HMI tags "Sim Stations"
   "HMI Data: Warehouse HMI_simStations_down" : Push Button Data = PLC "HMI Data: Warehouse HMI".simStations.down, 100 ms
   "HMI Data: Warehouse HMI_simStations_me{0}" : Station: Sim Data = PLC "HMI Data: Warehouse HMI".simStations.me[0] AT %DB1.DBX0.0, 100 ms
   "HMI Data: Warehouse HMI_simStations_me{1}" : Station: Sim Data = PLC "HMI Data: Warehouse HMI".simStations.me[1], 100 ms
   "HMI Data: Warehouse HMI_simStations_me{10}" : Station: Sim Data = PLC "HMI Data: Warehouse HMI".simStations.me[10], 100 ms
   "HMI Data: Warehouse HMI_simStations_me{11}" : Station: Sim Data = PLC "HMI Data: Warehouse HMI".simStations.me[11], 100 ms
   "HMI Data: Warehouse HMI_simStations_me{2}" : Station: Sim Data = PLC "HMI Data: Warehouse HMI".simStations.me[2], 100 ms
   "HMI Data: Warehouse HMI_simStations_me{3}" : Station: Sim Data = PLC "HMI Data: Warehouse HMI".simStations.me[3], 100 ms
   "HMI Data: Warehouse HMI_simStations_me{4}" : Station: Sim Data = PLC "HMI Data: Warehouse HMI".simStations.me[4], 100 ms
   "HMI Data: Warehouse HMI_simStations_me{5}" : Station: Sim Data = PLC "HMI Data: Warehouse HMI".simStations.me[5], 100 ms
   "HMI Data: Warehouse HMI_simStations_me{6}" : Station: Sim Data = PLC "HMI Data: Warehouse HMI".simStations.me[6], 100 ms
   "HMI Data: Warehouse HMI_simStations_me{7}" : Station: Sim Data = PLC "HMI Data: Warehouse HMI".simStations.me[7], 100 ms
   "HMI Data: Warehouse HMI_simStations_me{8}" : Station: Sim Data = PLC "HMI Data: Warehouse HMI".simStations.me[8], 100 ms
   "HMI Data: Warehouse HMI_simStations_me{9}" : Station: Sim Data = PLC "HMI Data: Warehouse HMI".simStations.me[9], 100 ms
   "HMI Data: Warehouse HMI_simStations_up" : Push Button Data = PLC "HMI Data: Warehouse HMI".simStations.up, 100 ms

HMI tags "Settings: Interface"
   "HMI Data: Warehouse HMI_settings_assign" : Push Button Data = PLC "HMI Data: Warehouse HMI".settings.assign, 100 ms
   "HMI Data: Warehouse HMI_settings_partNumber" : Part_Number_Double.UDT = PLC "HMI Data: Warehouse HMI".settings.partNumber, 100 ms
   "HMI Data: Warehouse HMI_settings_critical" : IO Field Data: Label with Data = PLC "HMI Data: Warehouse HMI".settings.critical, 100 ms
   "HMI Data: Warehouse HMI_settings_total" : IO Field Data: Label with Data = PLC "HMI Data: Warehouse HMI".settings.total, 100 ms
   "HMI Data: Warehouse HMI_settings_dropzone" : IO Field Data: Label with Data = PLC "HMI Data: Warehouse HMI".settings.dropzone, 100 ms
   "HMI Data: Warehouse HMI_settings_line" : IO Field Data: Label with Data = PLC "HMI Data: Warehouse HMI".settings.line, 100 ms
   "HMI Data: Warehouse HMI_settings_selectButton" : Push Button Data = PLC "HMI Data: Warehouse HMI".settings.selectButton, 100 ms
   "HMI Data: Warehouse HMI_settings_selectWip" : Push Button Data = PLC "HMI Data: Warehouse HMI".settings.selectWip, 100 ms
   "HMI Data: Warehouse HMI_settings_selectStation" : Push Button Data = PLC "HMI Data: Warehouse HMI".settings.selectStation, 100 ms
   "HMI Data: Warehouse HMI_settings_stnTableNavBar_hmi" : Nav Bar Data: HMI = PLC "HMI Data: Warehouse HMI".settings.stnTableNavBar.hmi AT %DB1.DBW0, 100 ms

HMI tags "Settings: Feedback"
   "HMI Data: Warehouse HMI_settings_stationRows{0}" : Settings Station Row Data = PLC "HMI Data: Warehouse HMI".settings.stationRows[0], 100 ms
   "HMI Data: Warehouse HMI_settings_stationRows{1}" : Settings Station Row Data = PLC "HMI Data: Warehouse HMI".settings.stationRows[1], 100 ms
   "HMI Data: Warehouse HMI_settings_stationRows{2}" : Settings Station Row Data = PLC "HMI Data: Warehouse HMI".settings.stationRows[2], 100 ms

graphic list "Vertical Table Nav Bar": 0 '100 x 100 Top'; 1 '100 x 100 Actuated Top'; 2 '100 x 100 Page Up'; 3 '100 x 100 Actuated Page Up'; 4 '100 x 100 Line Up'; 5 '100 x 100 Actuated Line Up'; 6 '100 x 100 Line Down'; 7 '100 x 100 Actuated Line Down'; 8 '100 x 100 Page Down'; 9 '100 x 100 Actuated Page Down'; 10 '100 x 100 Bottom'; 11 '100 x 100 Actuated Bottom'

screen "1 PART CALL" 1366x768
   on GenerateScreen: SetTag("HMI Data: Warehouse HMI_screenNumber", 1)
   Rectangle "Settings Tab Background" at 682,0 size 684x68
      Appearance <- "HMI Data: Warehouse HMI_screenNumber"
   Rectangle "Part Call Tab Background" at 0,0 size 685x68
      Appearance <- "HMI Data: Warehouse HMI_screenNumber"
   Rectangle "Settings Tab Border Hide" at 685,61 size 678x20
      Visibility <- "HMI Data: Warehouse HMI_screenNumber"
   Rectangle "Part Call Tab Border Hide" at 3,61 size 679x20
      Visibility <- "HMI Data: Warehouse HMI_screenNumber"
   Button "Settings Screen" at 683,0 size 683x68; TextOff 'SETTINGS'; Authorization "User administration"
      on Release: ActivateScreen("2 SETTINGS", 0)
   Button "Part Call Screen" at 0,0 size 683x68; TextOff 'PART CALL'
      on Release: ActivateScreen("1 PART CALL", 0)
   TextField "Header Line" at 32,112 size 216x53; Text 'LINE'
   TextField "Header Drop Zone" at 238,112 size 236x53; Text 'DROP ZONE'
   TextField "Header Part Number" at 474,112 size 648x53; Text 'PART NUMBER'
   TextField "Header Time" at 1112,112 size 222x53; Text 'TIME'
   ScreenModuleView "TableRow00" at 27,170 size 1312x52; ScreenModuleType ""
      Guid_{11997190-27688} <- "HMI Data: Warehouse HMI_partCall_row{0}"
      on Guid_{11997190-83214}: ActivateScreen("3 BARCODE", 0)
   ScreenModuleView "TableRow01" at 27,222 size 1312x52; ScreenModuleType ""
      Guid_{11997190-27688} <- "HMI Data: Warehouse HMI_partCall_row{1}"
      on Guid_{11997190-83214}: ActivateScreen("3 BARCODE", 0)
   ScreenModuleView "TableRow02" at 27,274 size 1312x52; ScreenModuleType ""
      Guid_{11997190-27688} <- "HMI Data: Warehouse HMI_partCall_row{2}"
      on Guid_{11997190-83214}: ActivateScreen("3 BARCODE", 0)
   ScreenModuleView "TableRow03" at 27,326 size 1312x52; ScreenModuleType ""
      Guid_{11997190-27688} <- "HMI Data: Warehouse HMI_partCall_row{3}"
      on Guid_{11997190-83214}: ActivateScreen("3 BARCODE", 0)
   ScreenModuleView "TableRow04" at 27,378 size 1312x52; ScreenModuleType ""
      Guid_{11997190-27688} <- "HMI Data: Warehouse HMI_partCall_row{4}"
      on Guid_{11997190-83214}: ActivateScreen("3 BARCODE", 0)
   ScreenModuleView "TableRow05" at 27,430 size 1312x52; ScreenModuleType ""
      Guid_{11997190-27688} <- "HMI Data: Warehouse HMI_partCall_row{5}"
      on Guid_{11997190-83214}: ActivateScreen("3 BARCODE", 0)
   ScreenModuleView "TableRow06" at 27,482 size 1312x52; ScreenModuleType ""
      Guid_{11997190-27688} <- "HMI Data: Warehouse HMI_partCall_row{6}"
      on Guid_{11997190-83214}: ActivateScreen("3 BARCODE", 0)
   ScreenModuleView "TableRow07" at 27,534 size 1312x52; ScreenModuleType ""
      Guid_{11997190-27688} <- "HMI Data: Warehouse HMI_partCall_row{7}"
      on Guid_{11997190-83214}: ActivateScreen("3 BARCODE", 0)
   ScreenModuleView "TableRow08" at 27,586 size 1312x52; ScreenModuleType ""
      Guid_{11997190-27688} <- "HMI Data: Warehouse HMI_partCall_row{8}"
      on Guid_{11997190-83214}: ActivateScreen("3 BARCODE", 0)
   ScreenModuleView "TableRow09" at 27,638 size 1312x52; ScreenModuleType ""
      Guid_{11997190-27688} <- "HMI Data: Warehouse HMI_partCall_row{9}"
      on Guid_{11997190-83214}: ActivateScreen("3 BARCODE", 0)
   ScreenModuleView "TableRow10" at 27,690 size 1312x52; ScreenModuleType ""
      Guid_{11997190-27688} <- "HMI Data: Warehouse HMI_partCall_row{10}"
      on Guid_{11997190-83214}: ActivateScreen("3 BARCODE", 0)

SlideinScreen "GraphX_Slidein_Bottom" 1366x80
   ScreenModuleView "Top" at 0,0 size 227x80; Guid_{11997190-63799} "Top"; ScreenModuleType ""
      Guid_{11997190-63779} <- "HMI Data: Warehouse HMI_tableNav_top"
   ScreenModuleView "Page Up" at 227,0 size 228x80; Guid_{11997190-63799} "pageUp"; ScreenModuleType ""
      Guid_{11997190-63779} <- "HMI Data: Warehouse HMI_tableNav_pageUp"
   ScreenModuleView "Line Up" at 455,0 size 228x80; Guid_{11997190-63799} "Up"; ScreenModuleType ""
      Guid_{11997190-63779} <- "HMI Data: Warehouse HMI_tableNav_lineUp"
   ScreenModuleView "Line Down" at 683,0 size 228x80; Guid_{11997190-63799} "Down"; ScreenModuleType ""
      Guid_{11997190-63779} <- "HMI Data: Warehouse HMI_tableNav_lineDown"
   ScreenModuleView "Page Down" at 911,0 size 228x80; Guid_{11997190-63799} "PageDown"; ScreenModuleType ""
      Guid_{11997190-63779} <- "HMI Data: Warehouse HMI_tableNav_pageDown"
   ScreenModuleView "Bottom" at 1138,0 size 228x80; Guid_{11997190-63799} "Bottom"; ScreenModuleType ""
      Guid_{11997190-63779} <- "HMI Data: Warehouse HMI_tableNav_bottom"
   TextField "Text field_1" at 0,0 size 1366x80; Text 'NOT USED'
      Visibility <- "HMI Data: Warehouse HMI_screenNumber"

SlideinScreen "GraphX_Slidein_Right" 449x768
   ScreenModuleView "Station Sim_1" at 5,5 size 106x232; ScreenModuleType ""
      Guid_{11997190-89108} <- "HMI Data: Warehouse HMI_simStations_me{0}"
   ScreenModuleView "Station Sim_2" at 116,5 size 106x232; ScreenModuleType ""
      Guid_{11997190-89108} <- "HMI Data: Warehouse HMI_simStations_me{1}"
   ScreenModuleView "Station Sim_3" at 227,5 size 106x232; ScreenModuleType ""
      Guid_{11997190-89108} <- "HMI Data: Warehouse HMI_simStations_me{2}"
   ScreenModuleView "Station Sim_4" at 338,5 size 106x232; ScreenModuleType ""
      Guid_{11997190-89108} <- "HMI Data: Warehouse HMI_simStations_me{3}"
   ScreenModuleView "Station Sim_5" at 5,242 size 106x232; ScreenModuleType ""
      Guid_{11997190-89108} <- "HMI Data: Warehouse HMI_simStations_me{4}"
   ScreenModuleView "Station Sim_6" at 5,479 size 106x232; ScreenModuleType ""
      Guid_{11997190-89108} <- "HMI Data: Warehouse HMI_simStations_me{8}"
   ScreenModuleView "Station Sim_7" at 116,242 size 106x232; ScreenModuleType ""
      Guid_{11997190-89108} <- "HMI Data: Warehouse HMI_simStations_me{5}"
   ScreenModuleView "Station Sim_8" at 227,242 size 106x232; ScreenModuleType ""
      Guid_{11997190-89108} <- "HMI Data: Warehouse HMI_simStations_me{6}"
   ScreenModuleView "Station Sim_9" at 338,242 size 106x232; ScreenModuleType ""
      Guid_{11997190-89108} <- "HMI Data: Warehouse HMI_simStations_me{7}"
   ScreenModuleView "Station Sim_10" at 116,479 size 106x232; ScreenModuleType ""
      Guid_{11997190-89108} <- "HMI Data: Warehouse HMI_simStations_me{9}"
   ScreenModuleView "Station Sim_11" at 227,478 size 106x232; ScreenModuleType ""
      Guid_{11997190-89108} <- "HMI Data: Warehouse HMI_simStations_me{10}"
   ScreenModuleView "Station Sim_12" at 338,477 size 106x232; ScreenModuleType ""
      Guid_{11997190-89108} <- "HMI Data: Warehouse HMI_simStations_me{11}"
   ScreenModuleView "PB: Graphic/Text List_1" at 5,716 size 65x45; Guid_{11997190-63799} "Up"; ScreenModuleType ""
      Guid_{11997190-63779} <- "HMI Data: Warehouse HMI_simStations_up"
   ScreenModuleView "PB: Graphic/Text List_2" at 379,716 size 65x45; Guid_{11997190-63799} "Down"; ScreenModuleType ""
      Guid_{11997190-63779} <- "HMI Data: Warehouse HMI_simStations_down"

screen "3 BARCODE" 1366x768
   on GenerateScreen: SetTag("HMI Data: Warehouse HMI_screenNumber", 3)
   Rectangle "Nav Panel 02" at 682,700 size 684x68
      Appearance <- "HMI Data: Warehouse HMI_screenNumber"
   Rectangle "Nav Panel 01" at 0,700 size 685x68
      Appearance <- "HMI Data: Warehouse HMI_screenNumber"
   Rectangle "Nav Panel 03 Top Border Hide" at 685,700 size 678x3
      Visibility <- "HMI Data: Warehouse HMI_screenNumber"
   Rectangle "Nav Panel 01 Top Border Hide" at 3,700 size 679x3
      Visibility <- "HMI Data: Warehouse HMI_screenNumber"
   Button "Settings Screen" at 683,700 size 683x68; TextOff 'SETTINGS'; Authorization "User administration"
      on Release: ActivateScreen("2 SETTINGS", 0)
   Button "Part Call Screen" at 0,700 size 683x68; TextOff 'PART CALL'
      on Release: ActivateScreen("1 PART CALL", 0)
   Button "btCancel" at 904,431 size 430x68; TextOff 'CANCEL'
      on Release: ActivateScreen("1 PART CALL", 0)
      on Press: function_b14e0dd5("animate_cancel", 0)
      Appearance <- "color_cancel"
   Button "btPartOrdered" at 32,431 size 430x68; TextOff 'ACKNOWLEDGED'
      on Release: SetBit("acknowledged"); ActivateScreen("1 PART CALL", 0)
      on Press: function_b14e0dd5("animate_acknowledged", 0)
      Appearance <- "color_acknowledged"
   TextField "tfBarcodeDisplay" at 32,220 size 1302x206; Text 'Text'
   TextField "tfPartNumberDisplay" at 32,160 size 1302x53; Text 'BARCODE FOR PART NUMBER'
   Button "btPartOrdered_1" at 468,431 size 430x68; TextOff 'ORDERED'
      on Release: SetBit("ordered"); ActivateScreen("1 PART CALL", 0)
      on Press: function_b14e0dd5("animate_ordered", 0)
      Appearance <- "color_ordered"

PopupScreen "KP8 Comm Status" 438x720
   ScreenModuleView "Station: KP8_1" at 5,5 size 428x710; ScreenModuleType ""
      Guid_{11997190-107144} <- "HMI Data: Warehouse HMI_networkHealth_kp8PopUp"
      on Guid_{11997190-107182}: function_efd93a16("KP8 Comm Status", 0, 0, -1, -1, 1)

PopupScreen "ET200SP Comm Status" 613x720
   ScreenModuleView "Station: ET200SP_1" at 5,5 size 603x710; ScreenModuleType ""
      Guid_{11997190-102952} <- "HMI Data: Warehouse HMI_networkHealth_et200spPopUp"
      on Guid_{11997190-102950}: function_efd93a16("ET200SP Comm Status", 0, 0, -1, -1, 1)

screen "2 SETTINGS" 1366x768
   on GenerateScreen: SetTag("HMI Data: Warehouse HMI_screenNumber", 2)
   Rectangle "Part Call Nave Panel" at 0,0 size 455x68
      Appearance <- "HMI Data: Warehouse HMI_screenNumber"
   Rectangle "Settings Nav Panel" at 452,0 size 462x68
      Appearance <- "HMI Data: Warehouse HMI_screenNumber"
   Rectangle "Network Health Nav Panel" at 911,0 size 455x68
      Appearance <- "HMI Data: Warehouse HMI_screenNumber"
   Rectangle "Part Call Border Hide" at 3,60 size 449x17
      Visibility <- "HMI Data: Warehouse HMI_screenNumber"
   Rectangle "Settings Border Hide" at 455,60 size 456x18
      Visibility <- "HMI Data: Warehouse HMI_screenNumber"
   Rectangle "Network Health Border Hide" at 914,60 size 449x18
      Visibility <- "HMI Data: Warehouse HMI_screenNumber"
   Button "Part Call Screen" at 0,0 size 455x68; TextOff 'PART CALL'
      on Release: ActivateScreen("1 PART CALL", 0)
   Button "Settings Screen" at 455,0 size 460x68; TextOff 'SETTINGS'
      on Release: ActivateScreen("2 SETTINGS", 0)
   Button "Network Health Screen" at 914,0 size 452x68; TextOff 'NW HEALTH'
   ScreenModuleView "pbSelectStation" at 60,108 size 370x55; Guid_{11997190-63616} 'Select Station'; ScreenModuleType ""
      on Guid_{11997190-211461}: function_efd93a16("Select Station", 30, 78, 1, -1, 1)
      Guid_{11997190-63605} <- "HMI Data: Warehouse HMI_settings_selectStation"
   ScreenModuleView "pbSelectWIP" at 60,173 size 370x56; Guid_{11997190-63616} 'Select WIP'; ScreenModuleType ""
      on Guid_{11997190-211461}: function_efd93a16("Select WIP", 30, 78, 1, -1, 1)
      Guid_{11997190-63605} <- "HMI Data: Warehouse HMI_settings_selectWip"
   ScreenModuleView "pbSelectButton" at 60,239 size 370x55; Guid_{11997190-63616} 'Select Button'; ScreenModuleType ""
      on Guid_{11997190-211461}: function_efd93a16("Select Button", 30, 78, 1, -1, 1)
      Guid_{11997190-63605} <- "HMI Data: Warehouse HMI_settings_selectButton"
   ScreenModuleView "pbAssign" at 60,652 size 370x56; Guid_{11997190-63616} 'Assign'; ScreenModuleType ""
      Guid_{11997190-63605} <- "HMI Data: Warehouse HMI_settings_assign"
   ScreenModuleView "iofLine" at 60,290 size 178x111; Guid_{11997190-206093} 'Line:'; ScreenModuleType ""
      Guid_{11997190-63113} <- "HMI Data: Warehouse HMI_settings_line"
   ScreenModuleView "iofDropzone" at 252,290 size 178x111; Guid_{11997190-206093} 'Dropzone:'; ScreenModuleType ""
      Guid_{11997190-63113} <- "HMI Data: Warehouse HMI_settings_dropzone"
   ScreenModuleView "iofAllotted" at 60,405 size 178x111; Guid_{11997190-206093} 'Total:'; ScreenModuleType ""
      Guid_{11997190-63113} <- "HMI Data: Warehouse HMI_settings_total"
   ScreenModuleView "iofCritical" at 252,405 size 178x111; Guid_{11997190-206093} 'Critical:'; ScreenModuleType ""
      Guid_{11997190-63113} <- "HMI Data: Warehouse HMI_settings_critical"
   TextField "tfHeaderLine" at 520,108 size 135x40; Text 'LINE'
   TextField "tfHeaderDropzone" at 655,108 size 40x40; Text 'DZ'
   TextField "tfHeaderWIP" at 695,108 size 40x40; Text 'WIP'
   TextField "tfHeaderButtonNumber" at 735,108 size 40x40; Text 'BTN'
   TextField "tfHeaderTotal" at 775,108 size 80x40; Text 'TOTAL'
   TextField "tfHeaderCritical" at 855,108 size 80x40; Text 'CRITICAL'
   TextField "tfHeaderPartNumber" at 935,108 size 256x40; Text 'PART NUMBER'
   ScreenModuleView "Settings Station Row_1" at 520,158 size 671x180; ScreenModuleType ""
      Guid_{11997190-213063} <- "HMI Data: Warehouse HMI_settings_stationRows{0}"
   ScreenModuleView "Settings Station Row_2" at 520,343 size 671x180; ScreenModuleType ""
      Guid_{11997190-213063} <- "HMI Data: Warehouse HMI_settings_stationRows{1}"
   ScreenModuleView "Settings Station Row_3" at 520,528 size 671x180; ScreenModuleType ""
      Guid_{11997190-213063} <- "HMI Data: Warehouse HMI_settings_stationRows{2}"
   ScreenModuleView "Settings Vertical Table Navigation" at 1206,108 size 100x600; ScreenModuleType ""
      Guid_{11997190-209443} <- "HMI Data: Warehouse HMI_settings_stnTableNavBar_hmi"
   ScreenModuleView "Part_Number_Entry" at 60,526 size 370x111; ScreenModuleType ""
      Guid_{11997190-63113} <- "HMI Data: Warehouse HMI_settings_partNumber"

PopupScreen "Select Station" 430x660
   TextField "Text field_1" at 30,30 size 325x40; Text 'Select Station'
   ScreenModuleView "Horizontal Table Navigation_1" at 30,568 size 372x62; ScreenModuleType ""
      Guid_{11997190-209443} <- "HMI Data: Warehouse HMI_pop_up_select_stations_nav_bar_hmi"
   ScreenModuleView "PB: Dynamic Text Label_1" at 30,85 size 178x65; ScreenModuleType ""
      Guid_{11997190-211129} <- "HMI Data: Warehouse HMI_pop_up_select_stations_stn_select_btns{0}"
   ScreenModuleView "PB: Dynamic Text Label_2" at 222,85 size 178x65; ScreenModuleType ""
      Guid_{11997190-211129} <- "HMI Data: Warehouse HMI_pop_up_select_stations_stn_select_btns{1}"
   ScreenModuleView "PB: Dynamic Text Label_3" at 30,165 size 178x65; ScreenModuleType ""
      Guid_{11997190-211129} <- "HMI Data: Warehouse HMI_pop_up_select_stations_stn_select_btns{2}"
   ScreenModuleView "PB: Dynamic Text Label_4" at 222,165 size 178x65; ScreenModuleType ""
      Guid_{11997190-211129} <- "HMI Data: Warehouse HMI_pop_up_select_stations_stn_select_btns{3}"
   ScreenModuleView "PB: Dynamic Text Label_5" at 30,245 size 178x65; ScreenModuleType ""
      Guid_{11997190-211129} <- "HMI Data: Warehouse HMI_pop_up_select_stations_stn_select_btns{4}"
   ScreenModuleView "PB: Dynamic Text Label_6" at 222,245 size 178x65; ScreenModuleType ""
      Guid_{11997190-211129} <- "HMI Data: Warehouse HMI_pop_up_select_stations_stn_select_btns{5}"
   ScreenModuleView "PB: Dynamic Text Label_7" at 30,325 size 178x65; ScreenModuleType ""
      Guid_{11997190-211129} <- "HMI Data: Warehouse HMI_pop_up_select_stations_stn_select_btns{6}"
   ScreenModuleView "PB: Dynamic Text Label_8" at 222,325 size 178x65; ScreenModuleType ""
      Guid_{11997190-211129} <- "HMI Data: Warehouse HMI_pop_up_select_stations_stn_select_btns{7}"
   ScreenModuleView "PB: Dynamic Text Label_9" at 30,405 size 178x65; ScreenModuleType ""
      Guid_{11997190-211129} <- "HMI Data: Warehouse HMI_pop_up_select_stations_stn_select_btns{8}"
   ScreenModuleView "PB: Dynamic Text Label_10" at 222,405 size 178x65; ScreenModuleType ""
      Guid_{11997190-211129} <- "HMI Data: Warehouse HMI_pop_up_select_stations_stn_select_btns{9}"
   ScreenModuleView "PB: Dynamic Text Label_11" at 30,485 size 178x65; ScreenModuleType ""
      Guid_{11997190-211129} <- "HMI Data: Warehouse HMI_pop_up_select_stations_stn_select_btns{10}"
   ScreenModuleView "PB: Dynamic Text Label_12" at 222,485 size 178x65; ScreenModuleType ""
      Guid_{11997190-211129} <- "HMI Data: Warehouse HMI_pop_up_select_stations_stn_select_btns{11}"
   ScreenModuleView "Close Select Station" at 360,30 size 40x40; Guid_{11997190-63799} "40 x 40 white close icon"; ScreenModuleType ""
      on Guid_{11997190-218589}: function_efd93a16("Select Station", 0, 0, 0, -1, 1)
      Guid_{11997190-63779} <- "HMI Data: Warehouse HMI_pop_up_select_stations_close_screen"

PopupScreen "Select WIP" 430x660
   TextField "Text field_1" at 30,30 size 325x40; Text 'Select WIP'
   ScreenModuleView "Horizontal Table Navigation_1" at 30,568 size 372x62; ScreenModuleType ""
      Guid_{11997190-209443} <- "HMI Data: Warehouse HMI_pop_up_select_WIPs_nav_bar_hmi"
   ScreenModuleView "PB: Dynamic Text Label_1" at 30,85 size 370x60; ScreenModuleType ""; Guid_{11997190-238549} "FontList_C3282863596"
      Guid_{11997190-211129} <- "HMI Data: Warehouse HMI_pop_up_select_WIPs_select_wip_buttons{0}"
   ScreenModuleView "PB: Dynamic Text Label_3" at 30,150 size 370x60; ScreenModuleType ""; Guid_{11997190-238549} "FontList_C3282863596"
      Guid_{11997190-211129} <- "HMI Data: Warehouse HMI_pop_up_select_WIPs_select_wip_buttons{1}"
   ScreenModuleView "PB: Dynamic Text Label_5" at 30,215 size 370x60; ScreenModuleType ""; Guid_{11997190-238549} "FontList_C3282863596"
      Guid_{11997190-211129} <- "HMI Data: Warehouse HMI_pop_up_select_WIPs_select_wip_buttons{2}"
   ScreenModuleView "PB: Dynamic Text Label_7" at 30,280 size 370x60; ScreenModuleType ""; Guid_{11997190-238549} "FontList_C3282863596"
      Guid_{11997190-211129} <- "HMI Data: Warehouse HMI_pop_up_select_WIPs_select_wip_buttons{3}"
   ScreenModuleView "PB: Dynamic Text Label_9" at 30,345 size 370x60; ScreenModuleType ""; Guid_{11997190-238549} "FontList_C3282863596"
      Guid_{11997190-211129} <- "HMI Data: Warehouse HMI_pop_up_select_WIPs_select_wip_buttons{4}"
   ScreenModuleView "PB: Dynamic Text Label_11" at 30,410 size 370x60; ScreenModuleType ""; Guid_{11997190-238549} "FontList_C3282863596"
      Guid_{11997190-211129} <- "HMI Data: Warehouse HMI_pop_up_select_WIPs_select_wip_buttons{5}"
   ScreenModuleView "PB: Dynamic Text Label_2" at 30,477 size 370x60; ScreenModuleType ""; Guid_{11997190-238549} "FontList_C3282863596"
      Guid_{11997190-211129} <- "HMI Data: Warehouse HMI_pop_up_select_WIPs_select_wip_buttons{6}"
   ScreenModuleView "PB: Graphic/Text List_1" at 360,30 size 40x40; ScreenModuleType ""; Guid_{11997190-63799} "40 x 40 white close icon"
      Guid_{11997190-63779} <- "HMI Data: Warehouse HMI_pop_up_select_WIPs_close_screen"
      on Guid_{11997190-218589}: function_efd93a16("Select WIP", 0, 0, 0, -1, 1)

PopupScreen "Select Button" 430x660
   GraphicView "Graphic view_1" at 0,0 size 430x660; Picture "kp8 image"
   ScreenModuleView "B01" at 95,90 size 105x105; Guid_{11997190-63616} '1'; ScreenModuleType ""
      Guid_{11997190-63605} <- "HMI Data: Warehouse HMI_pop_up_select_buttons_buttons{0}"
   ScreenModuleView "B02" at 228,90 size 105x105; Guid_{11997190-63616} '2'; ScreenModuleType ""
      Guid_{11997190-63605} <- "HMI Data: Warehouse HMI_pop_up_select_buttons_buttons{1}"
   ScreenModuleView "B03" at 95,213 size 105x105; Guid_{11997190-63616} '3'; ScreenModuleType ""
      Guid_{11997190-63605} <- "HMI Data: Warehouse HMI_pop_up_select_buttons_buttons{2}"
   ScreenModuleView "B05" at 95,336 size 105x105; Guid_{11997190-63616} '5'; ScreenModuleType ""
      Guid_{11997190-63605} <- "HMI Data: Warehouse HMI_pop_up_select_buttons_buttons{4}"
   ScreenModuleView "B07" at 95,459 size 105x105; Guid_{11997190-63616} '7'; ScreenModuleType ""
      Guid_{11997190-63605} <- "HMI Data: Warehouse HMI_pop_up_select_buttons_buttons{6}"
   ScreenModuleView "B04" at 228,213 size 105x105; Guid_{11997190-63616} '4'; ScreenModuleType ""
      Guid_{11997190-63605} <- "HMI Data: Warehouse HMI_pop_up_select_buttons_buttons{3}"
   ScreenModuleView "B06" at 228,336 size 105x105; Guid_{11997190-63616} '6'; ScreenModuleType ""
      Guid_{11997190-63605} <- "HMI Data: Warehouse HMI_pop_up_select_buttons_buttons{5}"
   ScreenModuleView "B08" at 228,459 size 105x105; Guid_{11997190-63616} '8'; ScreenModuleType ""
      Guid_{11997190-63605} <- "HMI Data: Warehouse HMI_pop_up_select_buttons_buttons{7}"
   ScreenModuleView "pb_close_pop_up" at 375,15 size 40x40; ScreenModuleType ""; Guid_{11997190-63799} "40 x 40 white close icon"
      on Guid_{11997190-218589}: function_efd93a16("Select Button", 0, 0, 0, -1, 1)
      Guid_{11997190-63779} <- "HMI Data: Warehouse HMI_pop_up_select_buttons_close_screen"
*)

(* ===== HMI "HMI_RT_2" =====
connection "LED Board": ETHERNET, S7_1500_OMS

HMI tags "Default tag table"
   "Clock_0.5Hz" : Bool = PLC "Clock_0.5Hz" AT %M0.7, 100 ms
   "LED Sign_request_row{0}" : Table Row = PLC "LED Sign".request.row[0], 100 ms
   "LED Sign_request_row{1}" : Table Row = PLC "LED Sign".request.row[1], 100 ms
   "LED Sign_request_row{2}" : Table Row = PLC "LED Sign".request.row[2], 100 ms
   "LED Sign_request_row{3}" : Table Row = PLC "LED Sign".request.row[3], 100 ms
   "LED Sign_request_row{4}" : Table Row = PLC "LED Sign".request.row[4], 100 ms
   "LED Sign_request_row{5}" : Table Row = PLC "LED Sign".request.row[5], 100 ms
   "LED Sign_request_row{6}" : Table Row = PLC "LED Sign".request.row[6], 100 ms
   "LED Sign_request_row{7}" : Table Row = PLC "LED Sign".request.row[7], 100 ms
   "LED Sign_request_row{8}" : Table Row = PLC "LED Sign".request.row[8], 100 ms
   "LED Sign_request_row{9}" : Table Row = PLC "LED Sign".request.row[9], 100 ms
   "LED Sign_request_row{10}" : Table Row = PLC "LED Sign".request.row[10], 100 ms
   "LED Sign_request_row{11}" : Table Row = PLC "LED Sign".request.row[11], 100 ms

screen "1 PART CALL" 1024x768
   Rectangle "Connection Status" at 1,196 size 894x1
      Appearance <- "Clock_0.5Hz"
   ScreenModuleView "R0C0" at 6,9 size 440x28; ScreenModuleType ""
      Guid_{11997190-27688} <- "LED Sign_request_row{0}"
   ScreenModuleView "R1C0" at 6,39 size 440x28; ScreenModuleType ""
      Guid_{11997190-27688} <- "LED Sign_request_row{1}"
   ScreenModuleView "R2C0" at 6,69 size 440x28; ScreenModuleType ""
      Guid_{11997190-27688} <- "LED Sign_request_row{2}"
   ScreenModuleView "R3C0" at 6,99 size 440x28; ScreenModuleType ""
      Guid_{11997190-27688} <- "LED Sign_request_row{3}"
   ScreenModuleView "R4C0" at 6,128 size 440x28; ScreenModuleType ""
      Guid_{11997190-27688} <- "LED Sign_request_row{4}"
   ScreenModuleView "R5C0" at 6,158 size 440x28; ScreenModuleType ""
      Guid_{11997190-27688} <- "LED Sign_request_row{5}"
   ScreenModuleView "R0C1" at 455,9 size 438x28; ScreenModuleType ""
      Guid_{11997190-27688} <- "LED Sign_request_row{6}"
   ScreenModuleView "R1C1" at 455,39 size 438x28; ScreenModuleType ""
      Guid_{11997190-27688} <- "LED Sign_request_row{7}"
   ScreenModuleView "R2C1" at 454,69 size 440x28; ScreenModuleType ""
      Guid_{11997190-27688} <- "LED Sign_request_row{8}"
   ScreenModuleView "R3C1" at 454,99 size 440x28; ScreenModuleType ""
      Guid_{11997190-27688} <- "LED Sign_request_row{9}"
   ScreenModuleView "R4C1" at 454,128 size 440x28; ScreenModuleType ""
      Guid_{11997190-27688} <- "LED Sign_request_row{10}"
   ScreenModuleView "R5C1" at 454,158 size 440x28; ScreenModuleType ""
      Guid_{11997190-27688} <- "LED Sign_request_row{11}"
*)

(* ===== HMI "HMI_RT_1" =====
system functions are stored by id; their names below are inferred from use

ScreenModuleEditorView "Table Row" 1312x52
   TextField "tfLine" at 5,1 size 216x48; Text 'Text'
      Visibility <- "interface.tfLine.visibility"
      Appearance <- "interface.tfLine.animator"
   TextField "tfTime" at 1085,1 size 222x48; Text 'Text'
      Appearance <- "interface.tfTime.animator"
      Visibility <- "interface.tfTime.visibility"
   TextField "tfDropZone" at 211,1 size 236x48; Text 'Text'
      Appearance <- "interface.tfDropZone.animator"
      Visibility <- "interface.tfDropZone.visibility"
   TextField "tfPartNumber" at 445,1 size 650x48; Text 'Text'
      Appearance <- "interface.tfPartNumber.animator"
      Visibility <- "interface.tfPartNumber.visibility"
   Button "pbSelect" at 0,0 size 1312x52; TextOff 'Text'
      Visibility <- "interface.pbSelection.visibility"
      on Press: SetBit("interface.pbSelection.request")
      on Release: ResetBit("interface.pbSelection.request")
   Rectangle "rtBackground" at 0,0 size 1312x52
      Visibility <- "interface.rtBackground.visibility"
*)

(* ===== HMI "HMI_RT_1" =====
system functions are stored by id; their names below are inferred from use

ScreenModuleEditorView "Table Row" 1312x52
   TextField "tfLine" at 5,1 size 216x48; Text 'Text'
      Visibility <- "interface.tfLine.visibility"
      Appearance <- "interface.tfLine.animator"
   TextField "tfTime" at 1085,1 size 222x48; Text 'Text'
      Visibility <- "interface.tfTime.visibility"
      Appearance <- "interface.tfTime.animator"
   TextField "tfDropZone" at 211,1 size 236x48; Text 'Text'
      Visibility <- "interface.tfDropZone.visibility"
      Appearance <- "interface.tfDropZone.animator"
   TextField "tfPartNumber" at 445,1 size 650x48; Text 'Text'
      Visibility <- "interface.tfPartNumber.visibility"
      Appearance <- "interface.tfPartNumber.animator"
   Button "pbSelect" at 0,0 size 1312x52; TextOff 'Text'
      on Release: ResetBit("interface.pbSelection.request")
      on Press: SetBit("interface.pbSelection.request")
      Visibility <- "interface.pbSelection.visibility"
   Rectangle "rtBackground" at 0,0 size 1312x52
      Visibility <- "interface.rtBackground.visibility"
*)

(* ===== HMI "HMI_RT_1" =====
system functions are stored by id; their names below are inferred from use

ScreenModuleEditorView "Table Row" 1312x52
   TextField "tfLine" at 5,1 size 216x48; Text 'Text'
      Visibility <- "interface.tfLine.visibility"
      Appearance <- "interface.tfLine.animator"
   TextField "tfTime" at 1085,1 size 222x48; Text 'Text'
      Visibility <- "interface.tfTime.visibility"
      Appearance <- "interface.tfTime.animator"
   TextField "tfDropZone" at 211,1 size 236x48; Text 'Text'
      Visibility <- "interface.tfDropZone.visibility"
      Appearance <- "interface.tfDropZone.animator"
   TextField "tfPartNumber" at 445,1 size 650x48; Text 'Text'
      Visibility <- "interface.tfPartNumber.visibility"
      Appearance <- "interface.tfPartNumber.animator"
   Button "pbSelect" at 0,0 size 1312x52; TextOff 'Text'
      on Release: ResetBit("interface.pbSelection.request")
      on Press: SetBit("interface.pbSelection.request")
      Visibility <- "interface.pbSelection.visibility"
   Rectangle "rtBackground" at 0,0 size 1312x52
      Visibility <- "interface.rtBackground.visibility"
*)

(* ===== HMI "HMI_RT_1" =====
system functions are stored by id; their names below are inferred from use

ScreenModuleEditorView "Table Row" 1312x52
   TextField "tfLine" at 5,1 size 216x48; Text 'Text'
      Visibility <- "interface.tfLine.visibility"
      Appearance <- "interface.tfLine.animator"
   TextField "tfTime" at 1085,1 size 222x48; Text 'Text'
      Visibility <- "interface.tfTime.visibility"
      Appearance <- "interface.tfTime.animator"
   TextField "tfDropZone" at 211,1 size 236x48; Text 'Text'
      Visibility <- "interface.tfDropZone.visibility"
      Appearance <- "interface.tfDropZone.animator"
   TextField "tfPartNumber" at 445,1 size 650x48; Text 'Text'
      Visibility <- "interface.tfPartNumber.visibility"
      Appearance <- "interface.tfPartNumber.animator"
   Button "pbSelect" at 0,0 size 1312x52; TextOff 'Text'
      on Release: ResetBit("interface.pbSelection.request")
      on Press: SetBit("interface.pbSelection.request")
      Visibility <- "interface.pbSelection.visibility"
   Rectangle "rtBackground" at 0,0 size 1312x52
      Visibility <- "interface.rtBackground.visibility"
*)

(* ===== HMI "HMI_RT_1" =====
system functions are stored by id; their names below are inferred from use

ScreenModuleEditorView "Table Row" 1312x52
   TextField "tfLine" at 5,1 size 216x48; Text 'Text'
      Visibility <- "interface.tfLine.visibility"
      Appearance <- "interface.tfLine.animator"
   TextField "tfTime" at 1085,1 size 222x48; Text 'Text'
      Visibility <- "interface.tfTime.visibility"
      Appearance <- "interface.tfTime.animator"
   TextField "tfDropZone" at 211,1 size 236x48; Text 'Text'
      Visibility <- "interface.tfDropZone.visibility"
      Appearance <- "interface.tfDropZone.animator"
   TextField "tfPartNumber" at 445,1 size 650x48; Text 'Text'
      Visibility <- "interface.tfPartNumber.visibility"
      Appearance <- "interface.tfPartNumber.animator"
   Button "pbSelect" at 0,0 size 1312x52; TextOff 'Text'
      on Release: ResetBit("interface.pbSelection.request")
      on Press: SetBit("interface.pbSelection.request")
      Visibility <- "interface.pbSelection.visibility"
   Rectangle "rtBackground" at 0,0 size 1312x52
      Visibility <- "interface.rtBackground.visibility"
*)

(* ===== HMI "HMI_RT_1" =====
system functions are stored by id; their names below are inferred from use

ScreenModuleEditorView "LED Row" 1312x52
   TextField "tfLine" at 5,1 size 216x48; Text 'Text'
      Visibility <- "interface.tfLine.visibility"
      Appearance <- "interface.tfLine.animator"
   TextField "tfTime" at 1085,1 size 222x48; Text 'Text'
      Visibility <- "interface.tfTime.visibility"
      Appearance <- "interface.tfTime.animator"
   TextField "tfDropZone" at 211,1 size 236x48; Text 'Text'
      Visibility <- "interface.tfDropZone.visibility"
      Appearance <- "interface.tfDropZone.animator"
   TextField "tfPartNumber" at 445,1 size 650x48; Text 'Text'
      Visibility <- "interface.tfPartNumber.visibility"
      Appearance <- "interface.tfPartNumber.animator"
   Button "pbSelect" at 0,0 size 1312x52; TextOff 'Text'
      on Release: ResetBit("interface.pbSelection.request")
      on Press: SetBit("interface.pbSelection.request")
      Visibility <- "interface.pbSelection.visibility"
   Rectangle "rtBackground" at 0,0 size 1312x52
      Visibility <- "interface.rtBackground.visibility"
*)

(* ===== HMI "HMI_RT_1" =====
system functions are stored by id; their names below are inferred from use

ScreenModuleEditorView "LED Row" 440x28
   TextField "tfLine" at 0,0 size 110x28; Text 'Text'
      Visibility <- "interface.tfLine.visibility"
      Appearance <- "interface.tfLine.animator"
   TextField "tfTime" at 349,0 size 91x28; Text 'Text'
      Visibility <- "interface.tfTime.visibility"
      Appearance <- "interface.tfTime.animator"
   TextField "tfDropZone" at 105,0 size 42x28; Text 'Text'
      Visibility <- "interface.tfDropZone.visibility"
      Appearance <- "interface.tfDropZone.animator"
   TextField "tfDLPartNumber" at 146,0 size 209x28; Text 'Text'
      Appearance <- "interface.tfPartNumber.animator"
      Visibility <- "interface.tfPartNumber.count"
   Button "pbSelect" at 0,0 size 440x28; TextOff 'Text'
      on Release: ResetBit("interface.pbSelection.request")
      on Press: SetBit("interface.pbSelection.request")
      Visibility <- "interface.pbSelection.visibility"
   Rectangle "rtBackground" at 0,0 size 440x28
      Visibility <- "interface.rtBackground.visibility"
   TextField "tfSLPartNumber" at 146,0 size 209x28; Text 'Text'
      Appearance <- "interface.tfPartNumber.animator"
      Visibility <- "interface.tfPartNumber.count"
*)

(* ===== HMI "HMI_RT_1" =====
system functions are stored by id; their names below are inferred from use

ScreenModuleEditorView "Table Row" 1312x52
   TextField "tfLine" at 5,1 size 216x48; Text 'Text'
      Visibility <- "interface.tfLine.visibility"
      Appearance <- "interface.tfLine.animator"
   TextField "tfTime" at 1085,1 size 222x48; Text 'Text'
      Visibility <- "interface.tfTime.visibility"
      Appearance <- "interface.tfTime.animator"
   TextField "tfDropZone" at 211,1 size 236x48; Text 'Text'
      Visibility <- "interface.tfDropZone.visibility"
      Appearance <- "interface.tfDropZone.animator"
   TextField "tfSLPartNumber" at 445,1 size 650x48; Text 'Text'
      Appearance <- "interface.tfPartNumber.animator"
      Visibility <- "interface.tfPartNumber.count"
   Button "pbSelect" at 0,0 size 1312x52; TextOff 'Text'
      on Release: ResetBit("interface.pbSelection.request")
      on Press: SetBit("interface.pbSelection.request")
      Visibility <- "interface.pbSelection.visibility"
   Rectangle "rtBackground" at 0,0 size 1312x52
      Visibility <- "interface.rtBackground.visibility"
   TextField "tfDLPartNumber" at 445,1 size 650x48; Text 'Text'
      Appearance <- "interface.tfPartNumber.animator"
      Visibility <- "interface.tfPartNumber.count"
*)

(* ===== HMI "HMI_RT_1" =====

ScreenModuleEditorView "LED Row" 440x28
   TextField "tfLine" at 0,0 size 110x28; Text 'Text'
      Visibility <- "interface.tfLine.visibility"
      Appearance <- "interface.tfLine.animator"
   TextField "tfTime" at 349,0 size 91x28; Text 'Text'
      Visibility <- "interface.tfTime.visibility"
      Appearance <- "interface.tfTime.animator"
   TextField "tfDropZone" at 105,0 size 42x28; Text 'Text'
      Visibility <- "interface.tfDropZone.visibility"
      Appearance <- "interface.tfDropZone.animator"
   TextField "tfSLPartNumber" at 146,0 size 209x28; Text 'Text'
      Visibility <- "interface.tfPartNumber.count"
      Appearance <- "interface.tfPartNumber.animator"
   TextField "tfDLPartNumber" at 146,0 size 209x28; Text 'Text'
      Visibility <- "interface.tfPartNumber.count"
      Appearance <- "interface.tfPartNumber.animator"
*)

(* ===== HMI "HMI_RT_1" =====
system functions are stored by id; their names below are inferred from use

ScreenModuleEditorView "Table Row" 1312x52
   TextField "tfLine" at 5,1 size 216x48; Text 'Text'
      Visibility <- "interface.tfLine.visibility"
      Appearance <- "interface.tfLine.animator"
   TextField "tfTime" at 1085,1 size 222x48; Text 'Text'
      Visibility <- "interface.tfTime.visibility"
      Appearance <- "interface.tfTime.animator"
   TextField "tfDropZone" at 211,1 size 236x48; Text 'Text'
      Visibility <- "interface.tfDropZone.visibility"
      Appearance <- "interface.tfDropZone.animator"
   TextField "tfSLPartNumber" at 445,1 size 650x48; Text 'Text'
      Visibility <- "interface.tfPartNumber.count"
      Appearance <- "interface.tfPartNumber.animator"
   Button "pbSelect" at 0,0 size 1312x52; TextOff 'Text'
      on Release: ResetBit("interface.pbSelection.request")
      on Press: SetBit("interface.pbSelection.request")
      Visibility <- "interface.pbSelection.visibility"
   Rectangle "rtBackground" at 0,0 size 1312x52
      Visibility <- "interface.rtBackground.visibility"
   TextField "tfDLPartNumber" at 445,1 size 650x48; Text 'Text'
      Visibility <- "interface.tfPartNumber.count"
      Appearance <- "interface.tfPartNumber.animator"
*)

(* ===== HMI "HMI_RT_1" =====
system functions are stored by id; their names below are inferred from use

ScreenModuleEditorView "PB: Station Select (Text Label)" 205x65
   Button "Station Select" at 0,0 size 205x65; TextOff 'Text'
      on Press: function_b14e0dd5("Interface.actuate", 0)
      Appearance <- "Interface.animate"
*)

(* ===== HMI "HMI_RT_1" =====
system functions are stored by id; their names below are inferred from use

ScreenModuleEditorView "PB: KP8 Button Select (Text Label)" 205x65
   Button "Station Select" at 0,0 size 205x65; TextOff 'Text'
      on Press: function_b14e0dd5("Interface.actuate", 0)
      Appearance <- "Interface.animate"
*)

(* ===== HMI "HMI_RT_1" =====
system functions are stored by id; their names below are inferred from use

ScreenModuleEditorView "PB: KP8 Button Select (Text Label)" 68x66
   Button "Station Select" at 0,0 size 68x66; TextOff 'Text'
      on Press: function_b14e0dd5("Interface.actuate", 0)
      Appearance <- "Interface.animate"
*)

(* ===== HMI "HMI_RT_1" =====
system functions are stored by id; their names below are inferred from use

ScreenModuleEditorView "PB: KP8 Stop Runtime (Text Label)" 68x66
   Button "Station Select" at 0,0 size 68x66; TextOff 'Text'
      on Press: function_b14e0dd5("Interface.actuate", 0)
      Appearance <- "Interface.animate"
*)

(* ===== HMI "HMI_RT_1" =====

ScreenModuleEditorView "PB: KP8 Stop Runtime (Text Label)" 68x66
   Button "Station Select" at 0,0 size 68x66; TextOff 'NOT USED'
      Appearance <- "Interface.animate"
*)

(* ===== HMI "HMI_RT_1" =====

ScreenModuleEditorView "PB: KP8 Stop Runtime (Text Label)" 68x66
   Button "Station Select" at 0,0 size 68x66; TextOff 'NOT USED'
      Appearance <- "Interface.animate"
*)

(* ===== HMI "HMI_RT_1" =====
system functions are stored by id; their names below are inferred from use

ScreenModuleEditorView "Station Assignment: Button Details" 513x74
   TextField "Button Label" at 0,0 size 75x74; Text 'Text'
      Appearance <- "Interface.label.animate"
      Visibility <- "Interface.label.animate"
   TextField "Critical Time" at 70,37 size 122x37; Text 'Text'
      Appearance <- "Interface.critical.animate"
      Visibility <- "Interface.critical.animate"
   TextField "Alloted Time" at 70,0 size 122x38; Text 'Text'
      Appearance <- "Interface.alloted.animate"
      Visibility <- "Interface.alloted.animate"
   TextField "Part Number" at 185,0 size 328x74; Text 'Text'
      Appearance <- "Interface.partNumber.animate"
      Visibility <- "Interface.partNumber.animate"
   Button "Select PB" at 0,0 size 513x74; TextOff 'Text'
      on Press: function_b14e0dd5("Interface.select.actuate", 0)
      Visibility <- "Interface.select.animate"
      ObjectEnable <- "Interface.select.animate"
*)

(* ===== HMI "HMI_RT_1" =====
system functions are stored by id; their names below are inferred from use

ScreenModuleEditorView "IO Field: Double Width: Stacked" 414x50
   IOField "PN Entry Field" at 0,0 size 414x50; FormatPattern ????????????????????????????????????????
      on OnFinishInput: SetBit("Interface.inputFinished")
      ObjectEnable <- "Interface.animate"
      Appearance <- "Interface.animate"
      ProcessValue <- "Interface.value"
*)

(* ===== HMI "HMI_RT_1" =====
system functions are stored by id; their names below are inferred from use

ScreenModuleEditorView "IO Field: Timer" 137x50
   IOField "Allotted Time Entry Field" at 0,0 size 137x50; FormatPattern ???????
      Appearance <- "Interface.animate"
      ObjectEnable <- "Interface.animate"
      on OnFinishInput: SetBit("Interface.inputFinished")
      ProcessValue <- "Interface.value"
*)

(* ===== HMI "HMI_RT_1" =====
system functions are stored by id; their names below are inferred from use

ScreenModuleEditorView "PB: Static Text Label" 274x45
   Button "Select All Stations" at 0,0 size 274x45; TextOff 'Text'
      on Press: function_b14e0dd5("Interface.actuate", 0)
      Appearance <- "Interface.animate"
*)

(* ===== HMI "HMI_RT_1" =====
system functions are stored by id; their names below are inferred from use

ScreenModuleEditorView "PB: Graphic/Text List" 65x45
   Button "Previous Station Group" at 0,0 size 65x45; TextOff 'Text'
      Visibility <- "Interface.animate"
      ObjectEnable <- "Interface.animate"
      Appearance <- "Interface.animate"
      on Press: SetBit("Interface.actuate")
*)

(* ===== HMI "HMI_RT_1" =====
system functions are stored by id; their names below are inferred from use

ScreenModuleEditorView "Line Label" 267x40
   IOField "Line" at 86,0 size 181x40; FormatPattern ?????????
      Appearance <- "interface.animate.ioField"
      ObjectEnable <- "interface.animate.ioField"
      Visibility <- "interface.animate.ioField"
      on OnFinishInput: SetBit("interface.inputFinished")
      ProcessValue <- "interface.value"
   TextField "Line Label" at 0,0 size 267x40; Text 'Line:'
      Appearance <- "interface.animate.bg"
      Visibility <- "interface.animate.bg"
*)

(* ===== HMI "HMI_RT_1" =====
system functions are stored by id; their names below are inferred from use

ScreenModuleEditorView "Drop Zone Label" 240x40
   IOField "Drop Zone Entry" at 171,0 size 69x40; FormatPattern ??
      Appearance <- "Interface.animate.ioField"
      ObjectEnable <- "Interface.animate.ioField"
      Visibility <- "Interface.animate.ioField"
      on OnFinishInput: SetBit("Interface.inputFinished")
      ProcessValue <- "Interface.value"
   TextField "Drop Zone Label" at 0,0 size 240x40; Text 'Drop Zone:'
      Appearance <- "Interface.animate.bg"
      Visibility <- "Interface.animate.bg"
*)

(* ===== HMI "HMI_RT_1" =====

ScreenModuleEditorView "PB: KP8 Reset Button (Text Label" 68x66
   Button "Station Select" at 0,0 size 68x66; TextOff 'NOT USED'
      Appearance <- "Interface.animate"
*)

(* ===== HMI "HMI_RT_1" =====

ScreenModuleEditorView "PB: KP8 Reset Button (Text Label" 68x66
   Button "Station Select" at 0,0 size 68x66; TextOff 'RESET SELECTED'
      Appearance <- "Interface.animate"
*)

(* ===== HMI "HMI_RT_1" =====

ScreenModuleEditorView "PB: KP8 Stop Runtime (Text Label)" 68x66
   Button "Station Select" at 0,0 size 68x66; TextOff 'STOP RUNTIME'
      Appearance <- "Interface.animate"
*)

(* ===== HMI "HMI_RT_1" =====
system functions are stored by id; their names below are inferred from use

ScreenModuleEditorView "PB: Graphic/Text List" 65x45
   Button "Previous Station Group" at 0,0 size 65x45; TextOff 'Text'
      on Press: SetBit("Interface.actuate")
      Visibility <- "Interface.animate"
      ObjectEnable <- "Interface.animate"
      Appearance <- "Interface.animate"
*)

(* ===== HMI "HMI_RT_1" =====
system functions are stored by id; their names below are inferred from use

ScreenModuleEditorView "PB: Static Text Label" 274x45
   Button "Select All Stations" at 0,0 size 274x45; TextOff 'Text'
      on Press: function_b14e0dd5("Interface.actuate", 0)
      Appearance <- "Interface.animate"
*)

(* ===== HMI "HMI_RT_1" =====
system functions are stored by id; their names below are inferred from use

ScreenModuleEditorView "PB: Static Text Label" 274x45
   Button "Select All Stations" at 0,0 size 274x45; TextOff 'Text'
      on Press: function_b14e0dd5("Interface.actuate", 0)
      Appearance <- "Interface.animate"
*)

(* ===== HMI "HMI_RT_1" =====
system functions are stored by id; their names below are inferred from use

ScreenModuleEditorView "PB: Graphic/Text List" 65x45
   Button "Previous Station Group" at 0,0 size 65x45; TextOff 'Text'
      on Press: SetBit("Interface.actuate")
      Visibility <- "Interface.animate"
      ObjectEnable <- "Interface.animate"
      Appearance <- "Interface.animate"
*)

(* ===== HMI "HMI_RT_1" =====
system functions are stored by id; their names below are inferred from use

ScreenModuleEditorView "PB: Station Select (Text Label)" 205x65
   Button "Station Select" at 0,0 size 205x65; TextOff 'Text'
      on Press: function_b14e0dd5("Interface.actuate", 0)
      Appearance <- "Interface.animate"
*)

(* ===== HMI "HMI_RT_1" =====
system functions are stored by id; their names below are inferred from use

ScreenModuleEditorView "PB: Graphic/Text List" 65x45
   Button "Previous Station Group" at 0,0 size 65x45; TextOff 'Text'
      on Press: function_b14e0dd5("Interface.actuate", 0)
      Visibility <- "Interface.animate"
      ObjectEnable <- "Interface.animate"
      Appearance <- "Interface.animate"
*)

(* ===== HMI "HMI_RT_1" =====
system functions are stored by id; their names below are inferred from use

ScreenModuleEditorView "Drop Zone Label" 240x40
   IOField "Drop Zone Entry" at 171,0 size 69x40; FormatPattern ??
      on OnFinishInput: SetBit("Interface.inputFinished")
      Appearance <- "Interface.animate.ioField"
      ObjectEnable <- "Interface.animate.ioField"
      Visibility <- "Interface.animate.ioField"
      ProcessValue <- "Interface.value"
   TextField "Drop Zone Label" at 0,0 size 240x40; Text 'Drop Zone:'
      Visibility <- "Interface.animate.bg"
      Appearance <- "Interface.animate.bg"
*)

(* ===== HMI "HMI_RT_1" =====
system functions are stored by id; their names below are inferred from use

ScreenModuleEditorView "IO Field: Double Width: Stacked" 414x50
   IOField "PN Entry Field" at 0,0 size 414x50; FormatPattern ????????????????????????????????????????
      on OnFinishInput: SetBit("Interface.inputFinished")
      Appearance <- "Interface.animate"
      ObjectEnable <- "Interface.animate"
      ProcessValue <- "Interface.value"
*)

(* ===== HMI "HMI_RT_1" =====
system functions are stored by id; their names below are inferred from use

ScreenModuleEditorView "IO Field: Timer" 137x50
   IOField "Allotted Time Entry Field" at 0,0 size 137x50; FormatPattern ???????
      on OnFinishInput: SetBit("Interface.inputFinished")
      Appearance <- "Interface.animate"
      ObjectEnable <- "Interface.animate"
      ProcessValue <- "Interface.value"
*)

(* ===== HMI "HMI_RT_1" =====